   "Carrier_72_G120DControlWord.14" AT %I3961.6 : Bool;   // Bit_14_DO0
   "Carrier_72_G120DControlWord.15" AT %I3961.7 : Bool;   // Bit_15_DO1
   "Carrier_72_G120DStatusWord" AT %IW3962 : Word;   // G120D_ZSW1_STATUS
   "Carrier_72_G120DStatusWord.0" AT %I3962.0 : Bool;   // Bit_00_READY_RUN
   "Carrier_72_G120DStatusWord.1" AT %I3962.1 : Bool;   // Bit_01_READY_ON
   "Carrier_72_G120DStatusWord.2" AT %I3962.2 : Bool;   // Bit_02_ENABLE
   "Carrier_72_G120DStatusWord.3" AT %I3962.3 : Bool;   // Bit_03_FAULT
   "Carrier_72_G120DStatusWord.4" AT %I3962.4 : Bool;   // Bit_04_OFF2
   "Carrier_72_G120DStatusWord.5" AT %I3962.5 : Bool;   // Bit_05_OFF3
   "Carrier_72_G120DStatusWord.6" AT %I3962.6 : Bool;   // Bit_06_LOCK_OUT
   "Carrier_72_G120DStatusWord.7" AT %I3962.7 : Bool;   // Bit_07_WARN
   "Carrier_72_G120DStatusWord.8" AT %I3963.0 : Bool;   // Bit_08_NO_DEVIATION
   "Carrier_72_G120DStatusWord.9" AT %I3963.1 : Bool;   // Bit_09_CONTR_PLC
   "Carrier_72_G120DStatusWord.10" AT %I3963.2 : Bool;   // Bit_10_F_MAX
   "Carrier_72_G120DStatusWord.11" AT %I3963.3 : Bool;   // Bit_11_LIMIT_REACHED
   "Carrier_72_G120DStatusWord.12" AT %I3963.4 : Bool;   // Bit_12_BRAKE_OPEN
   "Carrier_72_G120DStatusWord.13" AT %I3963.5 : Bool;   // Bit_13_NO_OVERTEMP
   "Carrier_72_G120DStatusWord.14" AT %I3963.6 : Bool;   // Bit_14_CW_CCW
   "Carrier_72_G120DStatusWord.15" AT %I3963.7 : Bool;   // Bit_15_OVERL
   "Carrier_72_Slot2_Input" AT %IW3964 : Word;   // SLOT 2 INPUT WORD
   "Carrier_72_CrashDetectSW" AT %I3964.0 : Bool;   // CRASH DETECT SW
   "Carrier_72_SpareSafetyInput(2_1)" AT %I3964.1 : Bool;   // SPARE SAFETY INPUT
   "Carrier_72_SpareSafetyInput(2_2)" AT %I3964.2 : Bool;   // SPARE SAFETY INPUT
   "Carrier_72_SpareSafetyInput(2_3)" AT %I3964.3 : Bool;   // SPARE SAFETY INPUT
   "Carrier_72_SpareSafetyInput(2_4)" AT %I3964.4 : Bool;   // SPARE SAFETY INPUT
   "Carrier_72_SpareSafetyInput(2_5)" AT %I3964.5 : Bool;   // SPARE SAFETY INPUT
   "Carrier_72_SpareSafetyInput(2_6)" AT %I3964.6 : Bool;   // SPARE SAFETY INPUT
   "Carrier_72_SpareSafetyInput(2_7)" AT %I3964.7 : Bool;   // SPARE SAFETY INPUT
   "Carrier_72_Slot3_SafetyOutput" AT %IW3965 : Word;   // SLOT 3 SAFETY OUTPUT WORD
   "Carrier_72_Crash_Detect_OK" AT %I3965.0 : Bool;   // CARRIER CRASH DETECT
   "Carrier_72_SpareSafetyOutput(3_1)" AT %I3965.1 : Bool;   // SPARE SAFETY OUTPUT
   "Carrier_72_SpareSafetyOutput(3_2)" AT %I3965.2 : Bool;   // SPARE SAFETY OUTPUT
   "Carrier_72_SpareSafetyOutput(3_3)" AT %I3965.3 : Bool;   // SPARE SAFETY OUTPUT
   "Carrier_72_SpareSafetyOutput(3_4)" AT %I3965.4 : Bool;   // SPARE SAFETY OUTPUT
   "Carrier_72_SpareSafetyOutput(3_5)" AT %I3965.5 : Bool;   // SPARE SAFETY OUTPUT
   "Carrier_72_SpareSafetyOutput(3_6)" AT %I3965.6 : Bool;   // SPARE SAFETY OUTPUT
   "Carrier_72_SpareSafetyOutput(3_7)" AT %I3965.7 : Bool;   // SPARE SAFETY OUTPUT
   "Carrier_72_Slot4_Input" AT %IW3966 : Word;   // SLOT 4 INPUT WORD
   "Carrier_72_480VPowerOn_MDCB1" AT %I3966.0 : Bool;   // 480 VAC POWER ON MDCB 1
   "Carrier_72_SpareInput(4_1)" AT %I3966.1 : Bool;   // SPARE INPUT
   "Carrier_72_SpareInput(4_2)" AT %I3966.2 : Bool;   // SPARE INPUT
   "Carrier_72_SitopSelectStatus" AT %I3966.3 : Bool;   // SITOP SELECT STATUS
   "Carrier_72_DCsupplyOnPSCB2" AT %I3966.4 : Bool;   // DC SUPPLY ON PSCB 2
   "Carrier_72_SpareInput(4_5)" AT %I3966.5 : Bool;   // SPARE INPUT
   "Carrier_72_SpareInput(4_6)" AT %I3966.6 : Bool;   // SPARE INPUT
   "Carrier_72_SpareInput(4_7)" AT %I3966.7 : Bool;   // SPARE INPUT
   "Carrier_72_PB1_ProdHoldLH" AT %I3967.0 : Bool;   // PB 1 PRODUCTION HOLD LH
   "Carrier_72_PB2_ResetLH" AT %I3967.1 : Bool;   // PB 2 RESET LH
   "Carrier_72_PB3_ProdHoldRH" AT %I3967.2 : Bool;   // PB 3 PRODUCTION HOLD RH
   "Carrier_72_PB4_ResetRH" AT %I3967.3 : Bool;   // PB 4 RESET RH
   "Carrier_72_SpareInput(4_14)" AT %I3967.4 : Bool;   // SPARE INPUT
   "Carrier_72_SpareInput(4_15)" AT %I3967.5 : Bool;   // SPARE INPUT
   "Carrier_72_SpareInput(4_16)" AT %I3967.6 : Bool;   // SPARE INPUT
   "Carrier_72_SpareInput(4_17)" AT %I3967.7 : Bool;   // SPARE INPUT
   "Carrier_72_Slot5_Output" AT %IW3968 : Word;   // SLOT 5 OUTPUT WORD
   "Carrier_72_IRD400_HMI_24VDC_ENABLE" AT %I3968.0 : Bool;   // IRD 400 PANEL HMI 24V DC POWER
   "Carrier_72_FaultLight_LH" AT %I3968.1 : Bool;   // FAULT LIGHT LH
   "Carrier_72_RunLight_LH" AT %I3968.2 : Bool;   // RUN LIGHT LH
   "Carrier_72_FaultLight_RH" AT %I3968.3 : Bool;   // FAULT LIGHT RH
   "Carrier_72_RunLight_RH" AT %I3968.4 : Bool;   // RUN LIGHT RH
   "Carrier_72_SpareOutput(5_5)" AT %I3968.5 : Bool;   // SPARE OUTPUT
   "Carrier_72_SpareOutput(5_6)" AT %I3968.6 : Bool;   // SPARE OUTPUT
   "Carrier_72_SpareOutput(5_7)" AT %I3968.7 : Bool;   // SPARE OUTPUT
   "Carrier_72_ActualSpeed" AT %IW3970 : Word;   // ACTUAL SPEED
   "Carrier_72_CarrierDriveAlarm" AT %IW3972 : Word;   // CARRIER DRIVE ALARM
   "Carrier_72_CarrierDriveWarning" AT %IW3974 : Word;   // CARRIER DRIVE WARNING
   "Carrier_73_Status" AT %IW4000 : Word;   // CARRIER STATUS WORD
   "Carrier_73_Status.0" AT %I4000.0 : Bool;   // HEARTBEAT
   "Carrier_73_Status.1" AT %I4000.1 : Bool;   // MANUAL
   "Carrier_73_Status.2" AT %I4000.2 : Bool;   // IN_AUTO
   "Carrier_73_Status.3" AT %I4000.3 : Bool;   // POSITIONING_COMPLETE
   "Carrier_73_Status.4" AT %I4000.4 : Bool;   // PRODUCTION HOLD
   "Carrier_73_Status.5" AT %I4000.5 : Bool;   // CARRIER MOVING FORWARD
   "Carrier_73_Status.6" AT %I4000.6 : Bool;   // CARRIER MOVING REVERSE
   "Carrier_73_Status.7" AT %I4000.7 : Bool;   // CARRIER FAULT
   "Carrier_73_Status.8" AT %I4001.0 : Bool;   // CRASH DETECT TRIPPED
   "Carrier_73_Status.9" AT %I4001.1 : Bool;
   "Carrier_73_Status.10" AT %I4001.2 : Bool;
   "Carrier_73_Status.11" AT %I4001.3 : Bool;
   "Carrier_73_Status.12" AT %I4001.4 : Bool;
   "Carrier_73_Status.13" AT %I4001.5 : Bool;
   "Carrier_73_Status.14" AT %I4001.6 : Bool;
   "Carrier_73_Status.15" AT %I4001.7 : Bool;
   "Carrier_73_SDCFaultCode" AT %IW4002 : Word;   // SDC FAULT CODE
   "Carrier_73_CarrierPosition" AT %ID4004 : DWord;   // CARRIER POSITION
   "Carrier_73_CarrierNumber" AT %IW4008 : Word;   // CARRIER NUMBER
   "Carrier_73_G120DControlWord" AT %IW4010 : Word;   // G120D_STW1_CONTROL
   "Carrier_73_G120DControlWord.0" AT %I4010.0 : Bool;   // Bit_00_ON
   "Carrier_73_G120DControlWord.1" AT %I4010.1 : Bool;   // Bit_01_AUS2_INH
   "Carrier_73_G120DControlWord.2" AT %I4010.2 : Bool;   // Bit_02_AUS3_STOP
   "Carrier_73_G120DControlWord.3" AT %I4010.3 : Bool;   // Bit_03_EN
   "Carrier_73_G120DControlWord.4" AT %I4010.4 : Bool;   // Bit_04_EN_RAMP
   "Carrier_73_G120DControlWord.5" AT %I4010.5 : Bool;   // Bit_05_START_RAMP
   "Carrier_73_G120DControlWord.6" AT %I4010.6 : Bool;   // Bit_06_SETPOINT
   "Carrier_73_G120DControlWord.7" AT %I4010.7 : Bool;   // Bit_07_RESET
   "Carrier_73_G120DControlWord.8" AT %I4011.0 : Bool;   // Bit_08_JOG_R
   "Carrier_73_G120DControlWord.9" AT %I4011.1 : Bool;   // Bit_09_JOG_L
   "Carrier_73_G120DControlWord.10" AT %I4011.2 : Bool;   // Bit_10_CONTR_PLC
   "Carrier_73_G120DControlWord.11" AT %I4011.3 : Bool;   // Bit_11_REVERSE
   "Carrier_73_G120DControlWord.12" AT %I4011.4 : Bool;   // Bit_12_BRAKE_RELEASE
   "Carrier_73_G120DControlWord.13" AT %I4011.5 : Bool;   // Bit_13_DDS
   "Carrier_73_G120DControlWord.14" AT %I4011.6 : Bool;   // Bit_14_DO0
   "Carrier_73_G120DControlWord.15" AT %I4011.7 : Bool;   // Bit_15_DO1
   "Carrier_73_G120DStatusWord" AT %IW4012 : Word;   // G120D_ZSW1_STATUS
   "Carrier_73_G120DStatusWord.0" AT %I4012.0 : Bool;   // Bit_00_READY_RUN
   "Carrier_73_G120DStatusWord.1" AT %I4012.1 : Bool;   // Bit_01_READY_ON
   "Carrier_73_G120DStatusWord.2" AT %I4012.2 : Bool;   // Bit_02_ENABLE
   "Carrier_73_G120DStatusWord.3" AT %I4012.3 : Bool;   // Bit_03_FAULT
   "Carrier_73_G120DStatusWord.4" AT %I4012.4 : Bool;   // Bit_04_OFF2
   "Carrier_73_G120DStatusWord.5" AT %I4012.5 : Bool;   // Bit_05_OFF3
   "Carrier_73_G120DStatusWord.6" AT %I4012.6 : Bool;   // Bit_06_LOCK_OUT
   "Carrier_73_G120DStatusWord.7" AT %I4012.7 : Bool;   // Bit_07_WARN
   "Carrier_73_G120DStatusWord.8" AT %I4013.0 : Bool;   // Bit_08_NO_DEVIATION
   "Carrier_73_G120DStatusWord.9" AT %I4013.1 : Bool;   // Bit_09_CONTR_PLC
   "Carrier_73_G120DStatusWord.10" AT %I4013.2 : Bool;   // Bit_10_F_MAX
   "Carrier_73_G120DStatusWord.11" AT %I4013.3 : Bool;   // Bit_11_LIMIT_REACHED
   "Carrier_73_G120DStatusWord.12" AT %I4013.4 : Bool;   // Bit_12_BRAKE_OPEN
   "Carrier_73_G120DStatusWord.13" AT %I4013.5 : Bool;   // Bit_13_NO_OVERTEMP
   "Carrier_73_G120DStatusWord.14" AT %I4013.6 : Bool;   // Bit_14_CW_CCW
   "Carrier_73_G120DStatusWord.15" AT %I4013.7 : Bool;   // Bit_15_OVERL
   "Carrier_73_Slot2_Input" AT %IW4014 : Word;   // SLOT 2 INPUT WORD
   "Carrier_73_CrashDetectSW" AT %I4014.0 : Bool;   // CRASH DETECT SW
   "Carrier_73_SpareSafetyInput(2_1)" AT %I4014.1 : Bool;   // SPARE SAFETY INPUT
   "Carrier_73_SpareSafetyInput(2_2)" AT %I4014.2 : Bool;   // SPARE SAFETY INPUT
   "Carrier_73_SpareSafetyInput(2_3)" AT %I4014.3 : Bool;   // SPARE SAFETY INPUT
   "Carrier_73_SpareSafetyInput(2_4)" AT %I4014.4 : Bool;   // SPARE SAFETY INPUT
   "Carrier_73_SpareSafetyInput(2_5)" AT %I4014.5 : Bool;   // SPARE SAFETY INPUT
   "Carrier_73_SpareSafetyInput(2_6)" AT %I4014.6 : Bool;   // SPARE SAFETY INPUT
   "Carrier_73_SpareSafetyInput(2_7)" AT %I4014.7 : Bool;   // SPARE SAFETY INPUT
   "Carrier_73_Slot3_SafetyOutput" AT %IW4015 : Word;   // SLOT 3 SAFETY OUTPUT WORD
   "Carrier_73_Crash_Detect_OK" AT %I4015.0 : Bool;   // CARRIER CRASH DETECT
   "Carrier_73_SpareSafetyOutput(3_1)" AT %I4015.1 : Bool;   // SPARE SAFETY OUTPUT
   "Carrier_73_SpareSafetyOutput(3_2)" AT %I4015.2 : Bool;   // SPARE SAFETY OUTPUT
   "Carrier_73_SpareSafetyOutput(3_3)" AT %I4015.3 : Bool;   // SPARE SAFETY OUTPUT
   "Carrier_73_SpareSafetyOutput(3_4)" AT %I4015.4 : Bool;   // SPARE SAFETY OUTPUT
   "Carrier_73_SpareSafetyOutput(3_5)" AT %I4015.5 : Bool;   // SPARE SAFETY OUTPUT
   "Carrier_73_SpareSafetyOutput(3_6)" AT %I4015.6 : Bool;   // SPARE SAFETY OUTPUT
   "Carrier_73_SpareSafetyOutput(3_7)" AT %I4015.7 : Bool;   // SPARE SAFETY OUTPUT
   "Carrier_73_Slot4_Input" AT %IW4016 : Word;   // SLOT 4 INPUT WORD
   "Carrier_73_480VPowerOn_MDCB1" AT %I4016.0 : Bool;   // 480 VAC POWER ON MDCB 1
   "Carrier_73_SpareInput(4_1)" AT %I4016.1 : Bool;   // SPARE INPUT
   "Carrier_73_SpareInput(4_2)" AT %I4016.2 : Bool;   // SPARE INPUT
   "Carrier_73_SitopSelectStatus" AT %I4016.3 : Bool;   // SITOP SELECT STATUS
   "Carrier_73_DCsupplyOnPSCB2" AT %I4016.4 : Bool;   // DC SUPPLY ON PSCB 2
   "Carrier_73_SpareInput(4_5)" AT %I4016.5 : Bool;   // SPARE INPUT
   "Carrier_73_SpareInput(4_6)" AT %I4016.6 : Bool;   // SPARE INPUT
   "Carrier_73_SpareInput(4_7)" AT %I4016.7 : Bool;   // SPARE INPUT
   "Carrier_73_PB1_ProdHoldLH" AT %I4017.0 : Bool;   // PB 1 PRODUCTION HOLD LH
   "Carrier_73_PB2_ResetLH" AT %I4017.1 : Bool;   // PB 2 RESET LH
   "Carrier_73_PB3_ProdHoldRH" AT %I4017.2 : Bool;   // PB 3 PRODUCTION HOLD RH
   "Carrier_73_PB4_ResetRH" AT %I4017.3 : Bool;   // PB 4 RESET RH
   "Carrier_73_SpareInput(4_14)" AT %I4017.4 : Bool;   // SPARE INPUT
   "Carrier_73_SpareInput(4_15)" AT %I4017.5 : Bool;   // SPARE INPUT
   "Carrier_73_SpareInput(4_16)" AT %I4017.6 : Bool;   // SPARE INPUT
   "Carrier_73_SpareInput(4_17)" AT %I4017.7 : Bool;   // SPARE INPUT
   "Carrier_73_Slot5_Output" AT %IW4018 : Word;   // SLOT 5 OUTPUT WORD
   "Carrier_73_IRD400_HMI_24VDC_ENABLE" AT %I4018.0 : Bool;   // IRD 400 PANEL HMI 24V DC POWER
   "Carrier_73_FaultLight_LH" AT %I4018.1 : Bool;   // FAULT LIGHT LH
   "Carrier_73_RunLight_LH" AT %I4018.2 : Bool;   // RUN LIGHT LH
   "Carrier_73_FaultLight_RH" AT %I4018.3 : Bool;   // FAULT LIGHT RH
   "Carrier_73_RunLight_RH" AT %I4018.4 : Bool;   // RUN LIGHT RH
   "Carrier_73_SpareOutput(5_5)" AT %I4018.5 : Bool;   // SPARE OUTPUT
   "Carrier_73_SpareOutput(5_6)" AT %I4018.6 : Bool;   // SPARE OUTPUT
   "Carrier_73_SpareOutput(5_7)" AT %I4018.7 : Bool;   // SPARE OUTPUT
   "Carrier_73_ActualSpeed" AT %IW4020 : Word;   // ACTUAL SPEED
   "Carrier_73_CarrierDriveAlarm" AT %IW4022 : Word;   // CARRIER DRIVE ALARM
   "Carrier_73_CarrierDriveWarning" AT %IW4024 : Word;   // CARRIER DRIVE WARNING
   "Carrier_74_Status" AT %IW4050 : Word;   // CARRIER STATUS WORD
   "Carrier_74_Status.0" AT %I4050.0 : Bool;   // HEARTBEAT
   "Carrier_74_Status.1" AT %I4050.1 : Bool;   // MANUAL
   "Carrier_74_Status.2" AT %I4050.2 : Bool;   // IN_AUTO
   "Carrier_74_Status.3" AT %I4050.3 : Bool;   // POSITIONING_COMPLETE
   "Carrier_74_Status.4" AT %I4050.4 : Bool;   // PRODUCTION HOLD
   "Carrier_74_Status.5" AT %I4050.5 : Bool;   // CARRIER MOVING FORWARD
   "Carrier_74_Status.6" AT %I4050.6 : Bool;   // CARRIER MOVING REVERSE
   "Carrier_74_Status.7" AT %I4050.7 : Bool;   // CARRIER FAULT
   "Carrier_74_Status.8" AT %I4051.0 : Bool;   // CRASH DETECT TRIPPED
   "Carrier_74_Status.9" AT %I4051.1 : Bool;
   "Carrier_74_Status.10" AT %I4051.2 : Bool;
   "Carrier_74_Status.11" AT %I4051.3 : Bool;
   "Carrier_74_Status.12" AT %I4051.4 : Bool;
   "Carrier_74_Status.13" AT %I4051.5 : Bool;
   "Carrier_74_Status.14" AT %I4051.6 : Bool;
   "Carrier_74_Status.15" AT %I4051.7 : Bool;
   "Carrier_74_SDCFaultCode" AT %IW4052 : Word;   // SDC FAULT CODE
   "Carrier_74_CarrierPosition" AT %ID4054 : DWord;   // CARRIER POSITION
   "Carrier_74_CarrierNumber" AT %IW4058 : Word;   // CARRIER NUMBER
   "Carrier_74_G120DControlWord" AT %IW4060 : Word;   // G120D_STW1_CONTROL
   "Carrier_74_G120DControlWord.0" AT %I4060.0 : Bool;   // Bit_00_ON
   "Carrier_74_G120DControlWord.1" AT %I4060.1 : Bool;   // Bit_01_AUS2_INH
   "Carrier_74_G120DControlWord.2" AT %I4060.2 : Bool;   // Bit_02_AUS3_STOP
   "Carrier_74_G120DControlWord.3" AT %I4060.3 : Bool;   // Bit_03_EN
   "Carrier_74_G120DControlWord.4" AT %I4060.4 : Bool;   // Bit_04_EN_RAMP
   "Carrier_74_G120DControlWord.5" AT %I4060.5 : Bool;   // Bit_05_START_RAMP
   "Carrier_74_G120DControlWord.6" AT %I4060.6 : Bool;   // Bit_06_SETPOINT
   "Carrier_74_G120DControlWord.7" AT %I4060.7 : Bool;   // Bit_07_RESET
   "Carrier_74_G120DControlWord.8" AT %I4061.0 : Bool;   // Bit_08_JOG_R
   "Carrier_74_G120DControlWord.9" AT %I4061.1 : Bool;   // Bit_09_JOG_L
   "Carrier_74_G120DControlWord.10" AT %I4061.2 : Bool;   // Bit_10_CONTR_PLC
   "Carrier_74_G120DControlWord.11" AT %I4061.3 : Bool;   // Bit_11_REVERSE
   "Carrier_74_G120DControlWord.12" AT %I4061.4 : Bool;   // Bit_12_BRAKE_RELEASE
   "Carrier_74_G120DControlWord.13" AT %I4061.5 : Bool;   // Bit_13_DDS
   "Carrier_74_G120DControlWord.14" AT %I4061.6 : Bool;   // Bit_14_DO0
   "Carrier_74_G120DControlWord.15" AT %I4061.7 : Bool;   // Bit_15_DO1
   "Carrier_74_G120DStatusWord" AT %IW4062 : Word;   // G120D_ZSW1_STATUS
   "Carrier_74_G120DStatusWord.0" AT %I4062.0 : Bool;   // Bit_00_READY_RUN
   "Carrier_74_G120DStatusWord.1" AT %I4062.1 : Bool;   // Bit_01_READY_ON
   "Carrier_74_G120DStatusWord.2" AT %I4062.2 : Bool;   // Bit_02_ENABLE
   "Carrier_74_G120DStatusWord.3" AT %I4062.3 : Bool;   // Bit_03_FAULT
   "Carrier_74_G120DStatusWord.4" AT %I4062.4 : Bool;   // Bit_04_OFF2
   "Carrier_74_G120DStatusWord.5" AT %I4062.5 : Bool;   // Bit_05_OFF3
   "Carrier_74_G120DStatusWord.6" AT %I4062.6 : Bool;   // Bit_06_LOCK_OUT
   "Carrier_74_G120DStatusWord.7" AT %I4062.7 : Bool;   // Bit_07_WARN
   "Carrier_74_G120DStatusWord.8" AT %I4063.0 : Bool;   // Bit_08_NO_DEVIATION
   "Carrier_74_G120DStatusWord.9" AT %I4063.1 : Bool;   // Bit_09_CONTR_PLC
   "Carrier_74_G120DStatusWord.10" AT %I4063.2 : Bool;   // Bit_10_F_MAX
   "Carrier_74_G120DStatusWord.11" AT %I4063.3 : Bool;   // Bit_11_LIMIT_REACHED
   "Carrier_74_G120DStatusWord.12" AT %I4063.4 : Bool;   // Bit_12_BRAKE_OPEN
   "Carrier_74_G120DStatusWord.13" AT %I4063.5 : Bool;   // Bit_13_NO_OVERTEMP
   "Carrier_74_G120DStatusWord.14" AT %I4063.6 : Bool;   // Bit_14_CW_CCW
   "Carrier_74_G120DStatusWord.15" AT %I4063.7 : Bool;   // Bit_15_OVERL
   "Carrier_74_Slot2_Input" AT %IW4064 : Word;   // SLOT 2 INPUT WORD
   "Carrier_74_CrashDetectSW" AT %I4064.0 : Bool;   // CRASH DETECT SW
   "Carrier_74_SpareSafetyInput(2_1)" AT %I4064.1 : Bool;   // SPARE SAFETY INPUT
   "Carrier_74_SpareSafetyInput(2_2)" AT %I4064.2 : Bool;   // SPARE SAFETY INPUT
   "Carrier_74_SpareSafetyInput(2_3)" AT %I4064.3 : Bool;   // SPARE SAFETY INPUT
   "Carrier_74_SpareSafetyInput(2_4)" AT %I4064.4 : Bool;   // SPARE SAFETY INPUT
   "Carrier_74_SpareSafetyInput(2_5)" AT %I4064.5 : Bool;   // SPARE SAFETY INPUT
   "Carrier_74_SpareSafetyInput(2_6)" AT %I4064.6 : Bool;   // SPARE SAFETY INPUT
   "Carrier_74_SpareSafetyInput(2_7)" AT %I4064.7 : Bool;   // SPARE SAFETY INPUT
   "Carrier_74_Slot3_SafetyOutput" AT %IW4065 : Word;   // SLOT 3 SAFETY OUTPUT WORD
   "Carrier_74_Crash_Detect_OK" AT %I4065.0 : Bool;   // CARRIER CRASH DETECT
   "Carrier_74_SpareSafetyOutput(3_1)" AT %I4065.1 : Bool;   // SPARE SAFETY OUTPUT
   "Carrier_74_SpareSafetyOutput(3_2)" AT %I4065.2 : Bool;   // SPARE SAFETY OUTPUT
   "Carrier_74_SpareSafetyOutput(3_3)" AT %I4065.3 : Bool;   // SPARE SAFETY OUTPUT
   "Carrier_74_SpareSafetyOutput(3_4)" AT %I4065.4 : Bool;   // SPARE SAFETY OUTPUT
   "Carrier_74_SpareSafetyOutput(3_5)" AT %I4065.5 : Bool;   // SPARE SAFETY OUTPUT
   "Carrier_74_SpareSafetyOutput(3_6)" AT %I4065.6 : Bool;   // SPARE SAFETY OUTPUT
   "Carrier_74_SpareSafetyOutput(3_7)" AT %I4065.7 : Bool;   // SPARE SAFETY OUTPUT
   "Carrier_74_Slot4_Input" AT %IW4066 : Word;   // SLOT 4 INPUT WORD
   "Carrier_74_480VPowerOn_MDCB1" AT %I4066.0 : Bool;   // 480 VAC POWER ON MDCB 1
   "Carrier_74_SpareInput(4_1)" AT %I4066.1 : Bool;   // SPARE INPUT
   "Carrier_74_SpareInput(4_2)" AT %I4066.2 : Bool;   // SPARE INPUT
   "Carrier_74_SitopSelectStatus" AT %I4066.3 : Bool;   // SITOP SELECT STATUS
   "Carrier_74_DCsupplyOnPSCB2" AT %I4066.4 : Bool;   // DC SUPPLY ON PSCB 2
   "Carrier_74_SpareInput(4_5)" AT %I4066.5 : Bool;   // SPARE INPUT
   "Carrier_74_SpareInput(4_6)" AT %I4066.6 : Bool;   // SPARE INPUT
   "Carrier_74_SpareInput(4_7)" AT %I4066.7 : Bool;   // SPARE INPUT
   "Carrier_74_PB1_ProdHoldLH" AT %I4067.0 : Bool;   // PB 1 PRODUCTION HOLD LH
   "Carrier_74_PB2_ResetLH" AT %I4067.1 : Bool;   // PB 2 RESET LH
   "Carrier_74_PB3_ProdHoldRH" AT %I4067.2 : Bool;   // PB 3 PRODUCTION HOLD RH
   "Carrier_74_PB4_ResetRH" AT %I4067.3 : Bool;   // PB 4 RESET RH
   "Carrier_74_SpareInput(4_14)" AT %I4067.4 : Bool;   // SPARE INPUT
   "Carrier_74_SpareInput(4_15)" AT %I4067.5 : Bool;   // SPARE INPUT
   "Carrier_74_SpareInput(4_16)" AT %I4067.6 : Bool;   // SPARE INPUT
   "Carrier_74_SpareInput(4_17)" AT %I4067.7 : Bool;   // SPARE INPUT
   "Carrier_74_Slot5_Output" AT %IW4068 : Word;   // SLOT 5 OUTPUT WORD
   "Carrier_74_IRD400_HMI_24VDC_ENABLE" AT %I4068.0 : Bool;   // IRD 400 PANEL HMI 24V DC POWER
   "Carrier_74_FaultLight_LH" AT %I4068.1 : Bool;   // FAULT LIGHT LH
   "Carrier_74_RunLight_LH" AT %I4068.2 : Bool;   // RUN LIGHT LH
   "Carrier_74_FaultLight_RH" AT %I4068.3 : Bool;   // FAULT LIGHT RH
   "Carrier_74_RunLight_RH" AT %I4068.4 : Bool;   // RUN LIGHT RH
   "Carrier_74_SpareOutput(5_5)" AT %I4068.5 : Bool;   // SPARE OUTPUT
   "Carrier_74_SpareOutput(5_6)" AT %I4068.6 : Bool;   // SPARE OUTPUT
   "Carrier_74_SpareOutput(5_7)" AT %I4068.7 : Bool;   // SPARE OUTPUT
   "Carrier_74_ActualSpeed" AT %IW4070 : Word;   // ACTUAL SPEED
   "Carrier_74_CarrierDriveAlarm" AT %IW4072 : Word;   // CARRIER DRIVE ALARM
   "Carrier_74_CarrierDriveWarning" AT %IW4074 : Word;   // CARRIER DRIVE WARNING
   "Carrier_75_Status" AT %IW4100 : Word;   // CARRIER STATUS WORD
   "Carrier_75_Status.0" AT %I4100.0 : Bool;   // HEARTBEAT
   "Carrier_75_Status.1" AT %I4100.1 : Bool;   // MANUAL
   "Carrier_75_Status.2" AT %I4100.2 : Bool;   // IN_AUTO
   "Carrier_75_Status.3" AT %I4100.3 : Bool;   // POSITIONING_COMPLETE
   "Carrier_75_Status.4" AT %I4100.4 : Bool;   // PRODUCTION HOLD
   "Carrier_75_Status.5" AT %I4100.5 : Bool;   // CARRIER MOVING FORWARD
   "Carrier_75_Status.6" AT %I4100.6 : Bool;   // CARRIER MOVING REVERSE
   "Carrier_75_Status.7" AT %I4100.7 : Bool;   // CARRIER FAULT
   "Carrier_75_Status.8" AT %I4101.0 : Bool;   // CRASH DETECT TRIPPED
   "Carrier_75_Status.9" AT %I4101.1 : Bool;
   "Carrier_75_Status.10" AT %I4101.2 : Bool;
   "Carrier_75_Status.11" AT %I4101.3 : Bool;
   "Carrier_75_Status.12" AT %I4101.4 : Bool;
   "Carrier_75_Status.13" AT %I4101.5 : Bool;
   "Carrier_75_Status.14" AT %I4101.6 : Bool;
   "Carrier_75_Status.15" AT %I4101.7 : Bool;
   "Carrier_75_SDCFaultCode" AT %IW4102 : Word;   // SDC FAULT CODE
   "Carrier_75_CarrierPosition" AT %ID4104 : DWord;   // CARRIER POSITION
   "Carrier_75_CarrierNumber" AT %IW4108 : Word;   // CARRIER NUMBER
   "Carrier_75_G120DControlWord" AT %IW4110 : Word;   // G120D_STW1_CONTROL
   "Carrier_75_G120DControlWord.0" AT %I4110.0 : Bool;   // Bit_00_ON
   "Carrier_75_G120DControlWord.1" AT %I4110.1 : Bool;   // Bit_01_AUS2_INH
   "Carrier_75_G120DControlWord.2" AT %I4110.2 : Bool;   // Bit_02_AUS3_STOP
   "Carrier_75_G120DControlWord.3" AT %I4110.3 : Bool;   // Bit_03_EN
   "Carrier_75_G120DControlWord.4" AT %I4110.4 : Bool;   // Bit_04_EN_RAMP
   "Carrier_75_G120DControlWord.5" AT %I4110.5 : Bool;   // Bit_05_START_RAMP
   "Carrier_75_G120DControlWord.6" AT %I4110.6 : Bool;   // Bit_06_SETPOINT
   "Carrier_75_G120DControlWord.7" AT %I4110.7 : Bool;   // Bit_07_RESET
   "Carrier_75_G120DControlWord.8" AT %I4111.0 : Bool;   // Bit_08_JOG_R
   "Carrier_75_G120DControlWord.9" AT %I4111.1 : Bool;   // Bit_09_JOG_L
   "Carrier_75_G120DControlWord.10" AT %I4111.2 : Bool;   // Bit_10_CONTR_PLC
   "Carrier_75_G120DControlWord.11" AT %I4111.3 : Bool;   // Bit_11_REVERSE
   "Carrier_75_G120DControlWord.12" AT %I4111.4 : Bool;   // Bit_12_BRAKE_RELEASE
   "Carrier_75_G120DControlWord.13" AT %I4111.5 : Bool;   // Bit_13_DDS
   "Carrier_75_G120DControlWord.14" AT %I4111.6 : Bool;   // Bit_14_DO0
   "Carrier_75_G120DControlWord.15" AT %I4111.7 : Bool;   // Bit_15_DO1
   "Carrier_75_G120DStatusWord" AT %IW4112 : Word;   // G120D_ZSW1_STATUS
   "Carrier_75_G120DStatusWord.0" AT %I4112.0 : Bool;   // Bit_00_READY_RUN
   "Carrier_75_G120DStatusWord.1" AT %I4112.1 : Bool;   // Bit_01_READY_ON
   "Carrier_75_G120DStatusWord.2" AT %I4112.2 : Bool;   // Bit_02_ENABLE
   "Carrier_75_G120DStatusWord.3" AT %I4112.3 : Bool;   // Bit_03_FAULT
   "Carrier_75_G120DStatusWord.4" AT %I4112.4 : Bool;   // Bit_04_OFF2
   "Carrier_75_G120DStatusWord.5" AT %I4112.5 : Bool;   // Bit_05_OFF3
   "Carrier_75_G120DStatusWord.6" AT %I4112.6 : Bool;   // Bit_06_LOCK_OUT
   "Carrier_75_G120DStatusWord.7" AT %I4112.7 : Bool;   // Bit_07_WARN
   "Carrier_75_G120DStatusWord.8" AT %I4113.0 : Bool;   // Bit_08_NO_DEVIATION
   "Carrier_75_G120DStatusWord.9" AT %I4113.1 : Bool;   // Bit_09_CONTR_PLC
   "Carrier_75_G120DStatusWord.10" AT %I4113.2 : Bool;   // Bit_10_F_MAX
   "Carrier_75_G120DStatusWord.11" AT %I4113.3 : Bool;   // Bit_11_LIMIT_REACHED
   "Carrier_75_G120DStatusWord.12" AT %I4113.4 : Bool;   // Bit_12_BRAKE_OPEN
   "Carrier_75_G120DStatusWord.13" AT %I4113.5 : Bool;   // Bit_13_NO_OVERTEMP
   "Carrier_75_G120DStatusWord.14" AT %I4113.6 : Bool;   // Bit_14_CW_CCW
   "Carrier_75_G120DStatusWord.15" AT %I4113.7 : Bool;   // Bit_15_OVERL
   "Carrier_75_Slot2_Input" AT %IW4114 : Word;   // SLOT 2 INPUT WORD
   "Carrier_75_CrashDetectSW" AT %I4114.0 : Bool;   // CRASH DETECT SW
   "Carrier_75_SpareSafetyInput(2_1)" AT %I4114.1 : Bool;   // SPARE SAFETY INPUT
   "Carrier_75_SpareSafetyInput(2_2)" AT %I4114.2 : Bool;   // SPARE SAFETY INPUT
   "Carrier_75_SpareSafetyInput(2_3)" AT %I4114.3 : Bool;   // SPARE SAFETY INPUT
   "Carrier_75_SpareSafetyInput(2_4)" AT %I4114.4 : Bool;   // SPARE SAFETY INPUT
   "Carrier_75_SpareSafetyInput(2_5)" AT %I4114.5 : Bool;   // SPARE SAFETY INPUT
   "Carrier_75_SpareSafetyInput(2_6)" AT %I4114.6 : Bool;   // SPARE SAFETY INPUT
   "Carrier_75_SpareSafetyInput(2_7)" AT %I4114.7 : Bool;   // SPARE SAFETY INPUT
   "Carrier_75_Slot3_SafetyOutput" AT %IW4115 : Word;   // SLOT 3 SAFETY OUTPUT WORD
   "Carrier_75_Crash_Detect_OK" AT %I4115.0 : Bool;   // CARRIER CRASH DETECT
   "Carrier_75_SpareSafetyOutput(3_1)" AT %I4115.1 : Bool;   // SPARE SAFETY OUTPUT
   "Carrier_75_SpareSafetyOutput(3_2)" AT %I4115.2 : Bool;   // SPARE SAFETY OUTPUT
   "Carrier_75_SpareSafetyOutput(3_3)" AT %I4115.3 : Bool;   // SPARE SAFETY OUTPUT
   "Carrier_75_SpareSafetyOutput(3_4)" AT %I4115.4 : Bool;   // SPARE SAFETY OUTPUT
   "Carrier_75_SpareSafetyOutput(3_5)" AT %I4115.5 : Bool;   // SPARE SAFETY OUTPUT
   "Carrier_75_SpareSafetyOutput(3_6)" AT %I4115.6 : Bool;   // SPARE SAFETY OUTPUT
   "Carrier_75_SpareSafetyOutput(3_7)" AT %I4115.7 : Bool;   // SPARE SAFETY OUTPUT
   "Carrier_75_Slot4_Input" AT %IW4116 : Word;   // SLOT 4 INPUT WORD
   "Carrier_75_480VPowerOn_MDCB1" AT %I4116.0 : Bool;   // 480 VAC POWER ON MDCB 1
   "Carrier_75_SpareInput(4_1)" AT %I4116.1 : Bool;   // SPARE INPUT
   "Carrier_75_SpareInput(4_2)" AT %I4116.2 : Bool;   // SPARE INPUT
   "Carrier_75_SitopSelectStatus" AT %I4116.3 : Bool;   // SITOP SELECT STATUS
   "Carrier_75_DCsupplyOnPSCB2" AT %I4116.4 : Bool;   // DC SUPPLY ON PSCB 2
   "Carrier_75_SpareInput(4_5)" AT %I4116.5 : Bool;   // SPARE INPUT
   "Carrier_75_SpareInput(4_6)" AT %I4116.6 : Bool;   // SPARE INPUT
   "Carrier_75_SpareInput(4_7)" AT %I4116.7 : Bool;   // SPARE INPUT
   "Carrier_75_PB1_ProdHoldLH" AT %I4117.0 : Bool;   // PB 1 PRODUCTION HOLD LH
   "Carrier_75_PB2_ResetLH" AT %I4117.1 : Bool;   // PB 2 RESET LH
   "Carrier_75_PB3_ProdHoldRH" AT %I4117.2 : Bool;   // PB 3 PRODUCTION HOLD RH
   "Carrier_75_PB4_ResetRH" AT %I4117.3 : Bool;   // PB 4 RESET RH
   "Carrier_75_SpareInput(4_14)" AT %I4117.4 : Bool;   // SPARE INPUT
   "Carrier_75_SpareInput(4_15)" AT %I4117.5 : Bool;   // SPARE INPUT
   "Carrier_75_SpareInput(4_16)" AT %I4117.6 : Bool;   // SPARE INPUT
   "Carrier_75_SpareInput(4_17)" AT %I4117.7 : Bool;   // SPARE INPUT
   "Carrier_75_Slot5_Output" AT %IW4118 : Word;   // SLOT 5 OUTPUT WORD
   "Carrier_75_IRD400_HMI_24VDC_ENABLE" AT %I4118.0 : Bool;   // IRD 400 PANEL HMI 24V DC POWER
   "Carrier_75_FaultLight_LH" AT %I4118.1 : Bool;   // FAULT LIGHT LH
   "Carrier_75_RunLight_LH" AT %I4118.2 : Bool;   // RUN LIGHT LH
   "Carrier_75_FaultLight_RH" AT %I4118.3 : Bool;   // FAULT LIGHT RH
   "Carrier_75_RunLight_RH" AT %I4118.4 : Bool;   // RUN LIGHT RH
   "Carrier_75_SpareOutput(5_5)" AT %I4118.5 : Bool;   // SPARE OUTPUT
   "Carrier_75_SpareOutput(5_6)" AT %I4118.6 : Bool;   // SPARE OUTPUT
   "Carrier_75_SpareOutput(5_7)" AT %I4118.7 : Bool;   // SPARE OUTPUT
   "Carrier_75_ActualSpeed" AT %IW4120 : Word;   // ACTUAL SPEED
   "Carrier_75_CarrierDriveAlarm" AT %IW4122 : Word;   // CARRIER DRIVE ALARM
   "Carrier_75_CarrierDriveWarning" AT %IW4124 : Word;   // CARRIER DRIVE WARNING
   "Carrier_76_Status" AT %IW4150 : Word;   // CARRIER STATUS WORD
   "Carrier_76_Status.0" AT %I4150.0 : Bool;   // HEARTBEAT
   "Carrier_76_Status.1" AT %I4150.1 : Bool;   // MANUAL
   "Carrier_76_Status.2" AT %I4150.2 : Bool;   // IN_AUTO
   "Carrier_76_Status.3" AT %I4150.3 : Bool;   // POSITIONING_COMPLETE
   "Carrier_76_Status.4" AT %I4150.4 : Bool;   // PRODUCTION HOLD
   "Carrier_76_Status.5" AT %I4150.5 : Bool;   // CARRIER MOVING FORWARD
   "Carrier_76_Status.6" AT %I4150.6 : Bool;   // CARRIER MOVING REVERSE
   "Carrier_76_Status.7" AT %I4150.7 : Bool;   // CARRIER FAULT
   "Carrier_76_Status.8" AT %I4151.0 : Bool;   // CRASH DETECT TRIPPED
   "Carrier_76_Status.9" AT %I4151.1 : Bool;
   "Carrier_76_Status.10" AT %I4151.2 : Bool;
   "Carrier_76_Status.11" AT %I4151.3 : Bool;
   "Carrier_76_Status.12" AT %I4151.4 : Bool;
   "Carrier_76_Status.13" AT %I4151.5 : Bool;
   "Carrier_76_Status.14" AT %I4151.6 : Bool;
   "Carrier_76_Status.15" AT %I4151.7 : Bool;
   "Carrier_76_SDCFaultCode" AT %IW4152 : Word;   // SDC FAULT CODE
   "Carrier_76_CarrierPosition" AT %ID4154 : DWord;   // CARRIER POSITION
   "Carrier_76_CarrierNumber" AT %IW4158 : Word;   // CARRIER NUMBER
   "Carrier_76_G120DControlWord" AT %IW4160 : Word;   // G120D_STW1_CONTROL
   "Carrier_76_G120DControlWord.0" AT %I4160.0 : Bool;   // Bit_00_ON
   "Carrier_76_G120DControlWord.1" AT %I4160.1 : Bool;   // Bit_01_AUS2_INH
   "Carrier_76_G120DControlWord.2" AT %I4160.2 : Bool;   // Bit_02_AUS3_STOP
   "Carrier_76_G120DControlWord.3" AT %I4160.3 : Bool;   // Bit_03_EN
   "Carrier_76_G120DControlWord.4" AT %I4160.4 : Bool;   // Bit_04_EN_RAMP
   "Carrier_76_G120DControlWord.5" AT %I4160.5 : Bool;   // Bit_05_START_RAMP
   "Carrier_76_G120DControlWord.6" AT %I4160.6 : Bool;   // Bit_06_SETPOINT
   "Carrier_76_G120DControlWord.7" AT %I4160.7 : Bool;   // Bit_07_RESET
   "Carrier_76_G120DControlWord.8" AT %I4161.0 : Bool;   // Bit_08_JOG_R
   "Carrier_76_G120DControlWord.9" AT %I4161.1 : Bool;   // Bit_09_JOG_L
   "Carrier_76_G120DControlWord.10" AT %I4161.2 : Bool;   // Bit_10_CONTR_PLC
   "Carrier_76_G120DControlWord.11" AT %I4161.3 : Bool;   // Bit_11_REVERSE
   "Carrier_76_G120DControlWord.12" AT %I4161.4 : Bool;   // Bit_12_BRAKE_RELEASE
   "Carrier_76_G120DControlWord.13" AT %I4161.5 : Bool;   // Bit_13_DDS
   "Carrier_76_G120DControlWord.14" AT %I4161.6 : Bool;   // Bit_14_DO0
   "Carrier_76_G120DControlWord.15" AT %I4161.7 : Bool;   // Bit_15_DO1
   "Carrier_76_G120DStatusWord" AT %IW4162 : Word;   // G120D_ZSW1_STATUS
   "Carrier_76_G120DStatusWord.0" AT %I4162.0 : Bool;   // Bit_00_READY_RUN
   "Carrier_76_G120DStatusWord.1" AT %I4162.1 : Bool;   // Bit_01_READY_ON
   "Carrier_76_G120DStatusWord.2" AT %I4162.2 : Bool;   // Bit_02_ENABLE
   "Carrier_76_G120DStatusWord.3" AT %I4162.3 : Bool;   // Bit_03_FAULT
   "Carrier_76_G120DStatusWord.4" AT %I4162.4 : Bool;   // Bit_04_OFF2
   "Carrier_76_G120DStatusWord.5" AT %I4162.5 : Bool;   // Bit_05_OFF3
   "Carrier_76_G120DStatusWord.6" AT %I4162.6 : Bool;   // Bit_06_LOCK_OUT
   "Carrier_76_G120DStatusWord.7" AT %I4162.7 : Bool;   // Bit_07_WARN
   "Carrier_76_G120DStatusWord.8" AT %I4163.0 : Bool;   // Bit_08_NO_DEVIATION
   "Carrier_76_G120DStatusWord.9" AT %I4163.1 : Bool;   // Bit_09_CONTR_PLC
   "Carrier_76_G120DStatusWord.10" AT %I4163.2 : Bool;   // Bit_10_F_MAX
   "Carrier_76_G120DStatusWord.11" AT %I4163.3 : Bool;   // Bit_11_LIMIT_REACHED
   "Carrier_76_G120DStatusWord.12" AT %I4163.4 : Bool;   // Bit_12_BRAKE_OPEN
   "Carrier_76_G120DStatusWord.13" AT %I4163.5 : Bool;   // Bit_13_NO_OVERTEMP
   "Carrier_76_G120DStatusWord.14" AT %I4163.6 : Bool;   // Bit_14_CW_CCW
   "Carrier_76_G120DStatusWord.15" AT %I4163.7 : Bool;   // Bit_15_OVERL
   "Carrier_76_Slot2_Input" AT %IW4164 : Word;   // SLOT 2 INPUT WORD
   "Carrier_76_CrashDetectSW" AT %I4164.0 : Bool;   // CRASH DETECT SW
   "Carrier_76_SpareSafetyInput(2_1)" AT %I4164.1 : Bool;   // SPARE SAFETY INPUT
   "Carrier_76_SpareSafetyInput(2_2)" AT %I4164.2 : Bool;   // SPARE SAFETY INPUT
   "Carrier_76_SpareSafetyInput(2_3)" AT %I4164.3 : Bool;   // SPARE SAFETY INPUT
   "Carrier_76_SpareSafetyInput(2_4)" AT %I4164.4 : Bool;   // SPARE SAFETY INPUT
   "Carrier_76_SpareSafetyInput(2_5)" AT %I4164.5 : Bool;   // SPARE SAFETY INPUT
   "Carrier_76_SpareSafetyInput(2_6)" AT %I4164.6 : Bool;   // SPARE SAFETY INPUT
   "Carrier_76_SpareSafetyInput(2_7)" AT %I4164.7 : Bool;   // SPARE SAFETY INPUT
   "Carrier_76_Slot3_SafetyOutput" AT %IW4165 : Word;   // SLOT 3 SAFETY OUTPUT WORD
   "Carrier_76_Crash_Detect_OK" AT %I4165.0 : Bool;   // CARRIER CRASH DETECT
   "Carrier_76_SpareSafetyOutput(3_1)" AT %I4165.1 : Bool;   // SPARE SAFETY OUTPUT
   "Carrier_76_SpareSafetyOutput(3_2)" AT %I4165.2 : Bool;   // SPARE SAFETY OUTPUT
   "Carrier_76_SpareSafetyOutput(3_3)" AT %I4165.3 : Bool;   // SPARE SAFETY OUTPUT
   "Carrier_76_SpareSafetyOutput(3_4)" AT %I4165.4 : Bool;   // SPARE SAFETY OUTPUT
   "Carrier_76_SpareSafetyOutput(3_5)" AT %I4165.5 : Bool;   // SPARE SAFETY OUTPUT
   "Carrier_76_SpareSafetyOutput(3_6)" AT %I4165.6 : Bool;   // SPARE SAFETY OUTPUT
   "Carrier_76_SpareSafetyOutput(3_7)" AT %I4165.7 : Bool;   // SPARE SAFETY OUTPUT
   "Carrier_76_Slot4_Input" AT %IW4166 : Word;   // SLOT 4 INPUT WORD
   "Carrier_76_480VPowerOn_MDCB1" AT %I4166.0 : Bool;   // 480 VAC POWER ON MDCB 1
   "Carrier_76_SpareInput(4_1)" AT %I4166.1 : Bool;   // SPARE INPUT
   "Carrier_76_SpareInput(4_2)" AT %I4166.2 : Bool;   // SPARE INPUT
   "Carrier_76_SitopSelectStatus" AT %I4166.3 : Bool;   // SITOP SELECT STATUS
   "Carrier_76_DCsupplyOnPSCB2" AT %I4166.4 : Bool;   // DC SUPPLY ON PSCB 2
   "Carrier_76_SpareInput(4_5)" AT %I4166.5 : Bool;   // SPARE INPUT
   "Carrier_76_SpareInput(4_6)" AT %I4166.6 : Bool;   // SPARE INPUT
   "Carrier_76_SpareInput(4_7)" AT %I4166.7 : Bool;   // SPARE INPUT
   "Carrier_76_PB1_ProdHoldLH" AT %I4167.0 : Bool;   // PB 1 PRODUCTION HOLD LH
   "Carrier_76_PB2_ResetLH" AT %I4167.1 : Bool;   // PB 2 RESET LH
   "Carrier_76_PB3_ProdHoldRH" AT %I4167.2 : Bool;   // PB 3 PRODUCTION HOLD RH
   "Carrier_76_PB4_ResetRH" AT %I4167.3 : Bool;   // PB 4 RESET RH
   "Carrier_76_SpareInput(4_14)" AT %I4167.4 : Bool;   // SPARE INPUT
   "Carrier_76_SpareInput(4_15)" AT %I4167.5 : Bool;   // SPARE INPUT
   "Carrier_76_SpareInput(4_16)" AT %I4167.6 : Bool;   // SPARE INPUT
   "Carrier_76_SpareInput(4_17)" AT %I4167.7 : Bool;   // SPARE INPUT